screen "0890_Consumption" 1280x800, template "Navigation"
   on GenerateScreen: SetTag("DB_Zaehler_Anzeige_ReadWriteDeviceNo", 1); "Consumtion"(); SetBit("DB_Zaehler_Anzeige_Read"); function_b431313b(2, U 1, N); SetTag("Recipe_Appearance_Control", 4)
   IOField "Cumulative" at 366,244 size 100x30; FormatPattern 999999
      ProcessValue <- "DB_Zaehler_Anzeige_Gesamt_Anzahl"
   IOField "I/O field_2" at 473,244 size 170x30; FormatPattern 999999.99
      ProcessValue <- "DB_Zaehler_Anzeige_Gesamt_Verbrauch_K1"
      Visibility <- "DB790_PlantParameter_AmountMeteringUnits"
   IOField "I/O field_3" at 650,244 size 170x30; FormatPattern 999999.99
      ProcessValue <- "DB_Zaehler_Anzeige_Gesamt_Verbrauch_K2"
      Visibility <- "DB790_PlantParameter_AmountMeteringUnits"
   Button "Button_1" at 960,145 size 181x53; TextOff 'Last Shift'; TextOn 'Actual Shift'; TextList "Consumtion_Button"
      on Press: InvertBit("DB_Zaehler_Anzeige_ViewPreShift"); SetBit("DB_Zaehler_Anzeige_Read")
      ProcessValue <- "DB_Zaehler_Anzeige_ViewPreShift"
   IOField "I/O field_4" at 650,328 size 170x30; FormatPattern 999999.99
      ProcessValue <- "DB_Zaehler_Anzeige_Counter{1}_Verbrauch_K2"
      Visibility <- "DB790_PlantParameter_AmountMeteringUnits"
   IOField "I/O field_5" at 650,367 size 170x30; FormatPattern 999999.99
      ProcessValue <- "DB_Zaehler_Anzeige_Counter{2}_Verbrauch_K2"
      Visibility <- "DB790_PlantParameter_AmountMeteringUnits"
   IOField "I/O field_6" at 650,405 size 170x30; FormatPattern 999999.99
      ProcessValue <- "DB_Zaehler_Anzeige_Counter{3}_Verbrauch_K2"
      Visibility <- "DB790_PlantParameter_AmountMeteringUnits"
   IOField "I/O field_7" at 650,444 size 170x30; FormatPattern 999999.99
      ProcessValue <- "DB_Zaehler_Anzeige_Counter{4}_Verbrauch_K2"
      Visibility <- "DB790_PlantParameter_AmountMeteringUnits"
   IOField "I/O field_8" at 650,483 size 170x30; FormatPattern 999999.99
      ProcessValue <- "DB_Zaehler_Anzeige_Counter{5}_Verbrauch_K2"
      Visibility <- "DB790_PlantParameter_AmountMeteringUnits"
   IOField "I/O field_9" at 650,521 size 170x30; FormatPattern 999999.99
      ProcessValue <- "DB_Zaehler_Anzeige_Counter{6}_Verbrauch_K2"
      Visibility <- "DB790_PlantParameter_AmountMeteringUnits"
   IOField "I/O field_10" at 650,560 size 170x30; FormatPattern 999999.99
      ProcessValue <- "DB_Zaehler_Anzeige_Counter{7}_Verbrauch_K2"
      Visibility <- "DB790_PlantParameter_AmountMeteringUnits"
   IOField "I/O field_11" at 650,598 size 170x30; FormatPattern 999999.99
      ProcessValue <- "DB_Zaehler_Anzeige_Counter{8}_Verbrauch_K2"
      Visibility <- "DB790_PlantParameter_AmountMeteringUnits"
   IOField "I/O field_12" at 650,638 size 170x30; FormatPattern 999999.99
      ProcessValue <- "DB_Zaehler_Anzeige_Counter{9}_Verbrauch_K2"
      Visibility <- "DB790_PlantParameter_AmountMeteringUnits"
   IOField "I/O field_13" at 650,675 size 170x30; FormatPattern 999999.99
      ProcessValue <- "DB_Zaehler_Anzeige_Counter{10}_Verbrauch_K2"
      Visibility <- "DB790_PlantParameter_AmountMeteringUnits"
   IOField "I/O field_14" at 473,328 size 170x30; FormatPattern 999999.99
      ProcessValue <- "DB_Zaehler_Anzeige_Counter{1}_Verbrauch_K1"
      Visibility <- "DB790_PlantParameter_AmountMeteringUnits"
   IOField "I/O field_15" at 473,367 size 170x30; FormatPattern 999999.99
      ProcessValue <- "DB_Zaehler_Anzeige_Counter{2}_Verbrauch_K1"
      Visibility <- "DB790_PlantParameter_AmountMeteringUnits"
   IOField "I/O field_16" at 473,405 size 170x30; FormatPattern 999999.99
      ProcessValue <- "DB_Zaehler_Anzeige_Counter{3}_Verbrauch_K1"
      Visibility <- "DB790_PlantParameter_AmountMeteringUnits"
   IOField "I/O field_17" at 473,444 size 170x30; FormatPattern 999999.99
      ProcessValue <- "DB_Zaehler_Anzeige_Counter{4}_Verbrauch_K1"
      Visibility <- "DB790_PlantParameter_AmountMeteringUnits"
   IOField "I/O field_18" at 473,483 size 170x30; FormatPattern 999999.99
      ProcessValue <- "DB_Zaehler_Anzeige_Counter{5}_Verbrauch_K1"
      Visibility <- "DB790_PlantParameter_AmountMeteringUnits"
   IOField "I/O field_19" at 473,521 size 170x30; FormatPattern 999999.99
      ProcessValue <- "DB_Zaehler_Anzeige_Counter{6}_Verbrauch_K1"
      Visibility <- "DB790_PlantParameter_AmountMeteringUnits"
   IOField "I/O field_20" at 473,560 size 170x30; FormatPattern 999999.99
      ProcessValue <- "DB_Zaehler_Anzeige_Counter{7}_Verbrauch_K1"
      Visibility <- "DB790_PlantParameter_AmountMeteringUnits"
   IOField "I/O field_21" at 473,598 size 170x30; FormatPattern 999999.99
      ProcessValue <- "DB_Zaehler_Anzeige_Counter{8}_Verbrauch_K1"
      Visibility <- "DB790_PlantParameter_AmountMeteringUnits"
   IOField "I/O field_22" at 473,638 size 170x30; FormatPattern 999999.99
      ProcessValue <- "DB_Zaehler_Anzeige_Counter{9}_Verbrauch_K1"
      Visibility <- "DB790_PlantParameter_AmountMeteringUnits"
   IOField "I/O field_23" at 473,675 size 170x30; FormatPattern 999999.99
      ProcessValue <- "DB_Zaehler_Anzeige_Counter{10}_Verbrauch_K1"
      Visibility <- "DB790_PlantParameter_AmountMeteringUnits"
   IOField "I/O field_24" at 366,327 size 100x30; FormatPattern 999999
      ProcessValue <- "DB_Zaehler_Anzeige_Counter{1}_Anzahl"
   IOField "I/O field_25" at 366,365 size 100x30; FormatPattern 999999
      ProcessValue <- "DB_Zaehler_Anzeige_Counter{2}_Anzahl"
   IOField "I/O field_26" at 366,405 size 100x30; FormatPattern 999999
      ProcessValue <- "DB_Zaehler_Anzeige_Counter{3}_Anzahl"
   IOField "I/O field_27" at 366,443 size 100x30; FormatPattern 999999
      ProcessValue <- "DB_Zaehler_Anzeige_Counter{4}_Anzahl"
   IOField "I/O field_28" at 366,481 size 100x30; FormatPattern 999999
      ProcessValue <- "DB_Zaehler_Anzeige_Counter{5}_Anzahl"
   IOField "I/O field_29" at 366,520 size 100x30; FormatPattern 999999
      ProcessValue <- "DB_Zaehler_Anzeige_Counter{6}_Anzahl"
   IOField "I/O field_30" at 366,558 size 100x30; FormatPattern 999999
      ProcessValue <- "DB_Zaehler_Anzeige_Counter{7}_Anzahl"
   IOField "I/O field_31" at 366,598 size 100x30; FormatPattern 999999
      ProcessValue <- "DB_Zaehler_Anzeige_Counter{8}_Anzahl"
   IOField "I/O field_32" at 366,637 size 100x30; FormatPattern 999999
      ProcessValue <- "DB_Zaehler_Anzeige_Counter{9}_Anzahl"
   IOField "I/O field_33" at 365,676 size 100x30; FormatPattern 999999
      ProcessValue <- "DB_Zaehler_Anzeige_Counter{10}_Anzahl"
   IOField "I/O field_34" at 178,326 size 180x30; FormatPattern ????????????????????????????????????????????????????????????????????????????????
      ProcessValue <- "Consumtion_Name_1"
   IOField "I/O field_35" at 178,364 size 180x30; FormatPattern ????????????????????????????????????????????????????????????????????????????????
      ProcessValue <- "Consumtion_Name_2"
   IOField "I/O field_36" at 178,404 size 180x30; FormatPattern ????????????????????????????????????????????????????????????????????????????????
      ProcessValue <- "Consumtion_Name_3"
   IOField "I/O field_37" at 178,441 size 180x30; FormatPattern ????????????????????????????????????????????????????????????????????????????????
      ProcessValue <- "Consumtion_Name_4"
   IOField "I/O field_38" at 178,480 size 180x30; FormatPattern ????????????????????????????????????????????????????????????????????????????????
      ProcessValue <- "Consumtion_Name_5"
   IOField "I/O field_39" at 178,519 size 180x30; FormatPattern ????????????????????????????????????????????????????????????????????????????????
      ProcessValue <- "Consumtion_Name_6"
   IOField "I/O field_40" at 178,558 size 180x30; FormatPattern ????????????????????????????????????????????????????????????????????????????????
      ProcessValue <- "Consumtion_Name_7"
   IOField "I/O field_41" at 178,597 size 180x30; FormatPattern ????????????????????????????????????????????????????????????????????????????????
      ProcessValue <- "Consumtion_Name_8"
   IOField "I/O field_42" at 178,636 size 180x30; FormatPattern ????????????????????????????????????????????????????????????????????????????????
      ProcessValue <- "Consumtion_Name_9"
   IOField "I/O field_43" at 178,676 size 180x30; FormatPattern ????????????????????????????????????????????????????????????????????????????????
      ProcessValue <- "Consumtion_Name_10"
   Button "Button_3" at 326,99 size 451x32; TextOff 'Consumption'
   Button "Button_2" at 293,154 size 313x35; TextOff '001--010'; TextList "Consumtion"
      ProcessValue <- "DB_Zaehler_Anzeige_ReadWriteDeviceNo"
   Button "Button_6" at 650,280 size 170x30; TextOff '[KG]'
      Visibility <- "DB790_PlantParameter_AmountMeteringUnits"
   Button "Button_7" at 366,280 size 100x30; TextOff 'Amount'
   Button "Button_8" at 178,244 size 180x30; TextOff 'Cumulative'
   Button "Button_9" at 178,280 size 180x30; TextOff 'Name'
   Button "Button_10" at 111,280 size 60x30; TextOff 'No'
   Button "Button_11" at 473,280 size 170x30; TextOff '[KG]'
      Visibility <- "DB790_PlantParameter_AmountMeteringUnits"
   Button "Button_12" at 121,326 size 50x30; TextOff '.'
   Button "Button_13" at 121,364 size 50x30; TextOff '.'
   Button "Button_14" at 121,404 size 50x30; TextOff '.'
   Button "Button_15" at 121,441 size 50x30; TextOff '.'
   Button "Button_16" at 121,480 size 50x30; TextOff '.'
   Button "Button_17" at 121,519 size 50x30; TextOff '.'
   Button "Button_18" at 121,558 size 50x30; TextOff '.'
   Button "Button_19" at 121,597 size 50x30; TextOff '.'
   Button "Button_20" at 121,636 size 50x30; TextOff '.'
   Button "Button_21" at 121,676 size 50x30; TextOff '.'
   Button "b_incress_consumtion" at 618,154 size 46x35; TextOff 'Text'; PictureOff "NEXT"
      on Click: "Consumtion_Increase"(); "Consumtion"(); SetBit("DB_Zaehler_Anzeige_Read"); function_dd21b452("Consumtion Name Multiplexing Control", 1)
   Button "b_Decres_consumtion" at 234,154 size 46x35; TextOff 'Text'; PictureOff "BEFORE"
      on Click: "Consumtiom_Decrease"(); "Consumtion"(); SetBit("DB_Zaehler_Anzeige_Read"); function_b9b71300("Consumtion Name Multiplexing Control", 1)
   IOField "I/O field_44" at 473,208 size 170x30; FormatPattern ????????????????????
      ProcessValue <- "DB753_MeteringPump_Pump{1}_Name"
      Appearance <- "DB702_Tank_Value_Tank{1}_Color"
      Visibility <- "DB790_PlantParameter_AmountMeteringUnits"
   IOField "I/O field_45" at 650,208 size 170x30; FormatPattern ????????????????????
      ProcessValue <- "DB753_MeteringPump_Pump{2}_Name"
      Appearance <- "DB702_Tank_Value_Tank{2}_Color"
      Visibility <- "DB790_PlantParameter_AmountMeteringUnits"
   IOField "I/O field_46" at 826,244 size 170x30; FormatPattern 999999.99
      ProcessValue <- "DB_Zaehler_Anzeige_Gesamt_Verbrauch_K3"
      Visibility <- "DB790_PlantParameter_AmountMeteringUnits"
   IOField "I/O field_47" at 1001,244 size 170x30; FormatPattern 999999.99
      ProcessValue <- "DB_Zaehler_Anzeige_Gesamt_Verbrauch_K4"
      Visibility <- "DB790_PlantParameter_AmountMeteringUnits"
   IOField "I/O field_48" at 1001,328 size 170x30; FormatPattern 999999.99
      ProcessValue <- "DB_Zaehler_Anzeige_Counter{1}_Verbrauch_K4"
      Visibility <- "DB790_PlantParameter_AmountMeteringUnits"
   IOField "I/O field_49" at 1001,367 size 170x30; FormatPattern 999999.99
      ProcessValue <- "DB_Zaehler_Anzeige_Counter{2}_Verbrauch_K4"
      Visibility <- "DB790_PlantParameter_AmountMeteringUnits"
   IOField "I/O field_50" at 1001,405 size 170x30; FormatPattern 999999.99
      ProcessValue <- "DB_Zaehler_Anzeige_Counter{3}_Verbrauch_K4"
      Visibility <- "DB790_PlantParameter_AmountMeteringUnits"
   IOField "I/O field_51" at 1001,444 size 170x30; FormatPattern 999999.99
      ProcessValue <- "DB_Zaehler_Anzeige_Counter{4}_Verbrauch_K4"
      Visibility <- "DB790_PlantParameter_AmountMeteringUnits"
   IOField "I/O field_52" at 1001,483 size 170x30; FormatPattern 999999.99
      ProcessValue <- "DB_Zaehler_Anzeige_Counter{5}_Verbrauch_K4"
      Visibility <- "DB790_PlantParameter_AmountMeteringUnits"
   IOField "I/O field_53" at 1001,521 size 170x30; FormatPattern 999999.99
      ProcessValue <- "DB_Zaehler_Anzeige_Counter{6}_Verbrauch_K4"
      Visibility <- "DB790_PlantParameter_AmountMeteringUnits"
   IOField "I/O field_54" at 1001,560 size 170x30; FormatPattern 999999.99
      ProcessValue <- "DB_Zaehler_Anzeige_Counter{7}_Verbrauch_K4"
      Visibility <- "DB790_PlantParameter_AmountMeteringUnits"
   IOField "I/O field_55" at 1001,598 size 170x30; FormatPattern 999999.99
      ProcessValue <- "DB_Zaehler_Anzeige_Counter{8}_Verbrauch_K4"
      Visibility <- "DB790_PlantParameter_AmountMeteringUnits"
   IOField "I/O field_56" at 1001,638 size 170x30; FormatPattern 999999.99
      ProcessValue <- "DB_Zaehler_Anzeige_Counter{9}_Verbrauch_K4"
      Visibility <- "DB790_PlantParameter_AmountMeteringUnits"
   IOField "I/O field_57" at 1001,675 size 170x30; FormatPattern 999999.99
      ProcessValue <- "DB_Zaehler_Anzeige_Counter{10}_Verbrauch_K4"
      Visibility <- "DB790_PlantParameter_AmountMeteringUnits"
   IOField "I/O field_58" at 826,328 size 170x30; FormatPattern 999999.99
      ProcessValue <- "DB_Zaehler_Anzeige_Counter{1}_Verbrauch_K3"
      Visibility <- "DB790_PlantParameter_AmountMeteringUnits"
   IOField "I/O field_59" at 826,367 size 170x30; FormatPattern 999999.99
      ProcessValue <- "DB_Zaehler_Anzeige_Counter{2}_Verbrauch_K3"
      Visibility <- "DB790_PlantParameter_AmountMeteringUnits"
   IOField "I/O field_60" at 826,405 size 170x30; FormatPattern 999999.99
      ProcessValue <- "DB_Zaehler_Anzeige_Counter{3}_Verbrauch_K3"
      Visibility <- "DB790_PlantParameter_AmountMeteringUnits"
   IOField "I/O field_61" at 826,444 size 170x30; FormatPattern 999999.99
      ProcessValue <- "DB_Zaehler_Anzeige_Counter{4}_Verbrauch_K3"
      Visibility <- "DB790_PlantParameter_AmountMeteringUnits"
   IOField "I/O field_62" at 826,483 size 170x30; FormatPattern 999999.99
      ProcessValue <- "DB_Zaehler_Anzeige_Counter{5}_Verbrauch_K3"
      Visibility <- "DB790_PlantParameter_AmountMeteringUnits"
   IOField "I/O field_63" at 826,521 size 170x30; FormatPattern 999999.99
      ProcessValue <- "DB_Zaehler_Anzeige_Counter{6}_Verbrauch_K3"
      Visibility <- "DB790_PlantParameter_AmountMeteringUnits"
   IOField "I/O field_64" at 826,560 size 170x30; FormatPattern 999999.99
      ProcessValue <- "DB_Zaehler_Anzeige_Counter{7}_Verbrauch_K3"
      Visibility <- "DB790_PlantParameter_AmountMeteringUnits"
   IOField "I/O field_65" at 826,598 size 170x30; FormatPattern 999999.99
      ProcessValue <- "DB_Zaehler_Anzeige_Counter{8}_Verbrauch_K3"
      Visibility <- "DB790_PlantParameter_AmountMeteringUnits"
   IOField "I/O field_66" at 826,638 size 170x30; FormatPattern 999999.99
      ProcessValue <- "DB_Zaehler_Anzeige_Counter{9}_Verbrauch_K3"
      Visibility <- "DB790_PlantParameter_AmountMeteringUnits"
   IOField "I/O field_67" at 826,675 size 170x30; FormatPattern 999999.99
      ProcessValue <- "DB_Zaehler_Anzeige_Counter{10}_Verbrauch_K3"
      Visibility <- "DB790_PlantParameter_AmountMeteringUnits"
   Button "Button_4" at 1001,280 size 170x30; TextOff '[KG]'
      Visibility <- "DB790_PlantParameter_AmountMeteringUnits"
   Button "Button_5" at 826,280 size 170x30; TextOff '[KG]'
      Visibility <- "DB790_PlantParameter_AmountMeteringUnits"
   IOField "I/O field_68" at 826,208 size 170x30; FormatPattern ????????????????????
      ProcessValue <- "DB753_MeteringPump_Pump{3}_Name"
      Visibility <- "DB790_PlantParameter_AmountMeteringUnits"
      Appearance <- "DB702_Tank_Value_Tank{3}_Color"
   IOField "I/O field_69" at 1001,208 size 170x30; FormatPattern ????????????????????
      ProcessValue <- "DB753_MeteringPump_Pump{4}_Name"
      Visibility <- "DB790_PlantParameter_AmountMeteringUnits"
      Appearance <- "DB702_Tank_Value_Tank{4}_Color"
   Button "b_ShifProto_ShotCounter_1" at 208,713 size 60x60; TextOff 'Shot Counter'; PictureList "ico_ShiftProtocol"
      ProcessValue <- "Recipe_Appearance_Control"
      Appearance <- "Recipe_Appearance_Control"
   Button "b_Shiftproto_shiftproto" at 208,713 size 60x60; TextOff 'Shift proto'
      on Click: ActivateScreen("0112_Shift protocol", 0); SetTag("Recipe_Appearance_Control", 2)
      Appearance <- "Recipe_Appearance_Control"
   Button "b_SC" at 478,713 size 60x60; TextOff 'Shot Counter'; PictureList "ico_ShotCounter"
      on Press: ActivateScreen("0891_Shotcounter MixingHead", 0); SetTag("Recipe_Appearance_Control", 5)
      Appearance <- "Recipe_Appearance_Control"
      ProcessValue <- "Recipe_Appearance_Control"
   Button "b_SC_1" at 478,713 size 60x60; TextOff 'Shot Counter'
      on Click: ActivateScreen("0891_Shotcounter MixingHead", 0); SetTag("Recipe_Appearance_Control", 5)
      Appearance <- "Recipe_Appearance_Control"
   Button "b_Shift_Plan" at 118,713 size 60x60; TextOff 'Shift Plan'; PictureList "ico_ShiftPlan"
      on Press: ActivateScreen("0113_SettingShiftPlan", 0); SetTag("Recipe_Appearance_Control", 1)
      Appearance <- "Recipe_Appearance_Control"
      ProcessValue <- "Recipe_Appearance_Control"
   Button "b_Shift_Plan_1" at 118,713 size 60x60; TextOff 'Shift Plan'
      on Click: "SettingShiftPlan"(); ActivateScreen("0113_SettingShiftPlan", 0); SetTag("Recipe_Appearance_Control", 1)
      Appearance <- "Recipe_Appearance_Control"
   Button "b_LS_Lastshot" at 298,713 size 60x60; TextOff 'Last Shot'; PictureList "ico_LastShot"
      on Press: ActivateScreen("0036_Last Shot", 0); SetTag("Recipe_Appearance_Control", 3)
      Appearance <- "Recipe_Appearance_Control"
      ProcessValue <- "Recipe_Appearance_Control"
   Button "b_LS_Lastshot_1" at 298,713 size 60x60; TextOff 'Last Shot'
      on Click: ActivateScreen("0036_Last Shot", 0); SetTag("Recipe_Appearance_Control", 3)
      Appearance <- "Recipe_Appearance_Control"
   Button "b_Consumtion" at 388,713 size 60x60; TextOff 'Consumtion / Consum'; PictureList "ico_consum"
      on Press: ActivateScreen("0890_Consumption", 0); SetTag("Recipe_Appearance_Control", 4)
      Appearance <- "Recipe_Appearance_Control"
      ProcessValue <- "Recipe_Appearance_Control"
   Button "b_Consumtion_1" at 388,713 size 60x60; TextOff 'Consumtion / Consum'
      on Click: ActivateScreen("0890_Consumption", 0); SetTag("Recipe_Appearance_Control", 4)
      Appearance <- "Recipe_Appearance_Control"

screen "0891_Shotcounter MixingHead" 1280x800, template "Navigation"
   on GenerateScreen: SetBit("DB_Zaehler_Anzeige_Read"); SetTag("Recipe_Appearance_Control", 5)
   IOField "I/O field_14" at 378,202 size 168x30; FormatPattern 9999999
      ProcessValue <- "DB_Zaehler_Anzeige_MH_Counter_ActualShift{1}"
      Visibility <- "DB790_PlantParameter_AmountMH"
   IOField "lastshift1" at 564,202 size 168x30; FormatPattern 9999999
      ProcessValue <- "DB_Zaehler_Anzeige_MH_Counter_PreShift{1}"
      Visibility <- "DB790_PlantParameter_AmountMH"
   IOField "I/O field_2" at 748,202 size 168x30; Authorization "User administration"; FormatPattern 9999999
      ProcessValue <- "DB_Zaehler_Anzeige_MH_Counter_Reset{1}"
      Visibility <- "DB790_PlantParameter_AmountMH"
   IOField "I/O field_3" at 933,202 size 168x30; FormatPattern 9999999
      ProcessValue <- "DB_Zaehler_Anzeige_MH_Counter_NonReset{1}"
      Visibility <- "DB790_PlantParameter_AmountMH"
   Button "Button_3" at 326,104 size 451x32; TextOff 'Shot counter Mixinghead'
   Button "Button_1" at 378,158 size 168x30; TextOff 'Actual Shift'
   Button "Button_2" at 564,158 size 168x30; TextOff 'Last Shift'
   Button "Button_4" at 748,158 size 168x30; TextOff 'Resetable'
   Button "Button_5" at 933,158 size 168x30; TextOff 'Cumulative'
   Button "Button_6" at 309,202 size 50x30; TextOff '1.'
      Visibility <- "DB790_PlantParameter_AmountMH"
   IOField "I/O field_4" at 378,245 size 168x30; FormatPattern 9999999
      ProcessValue <- "DB_Zaehler_Anzeige_MH_Counter_ActualShift{2}"
      Visibility <- "DB790_PlantParameter_AmountMH"
   IOField "I/O field_5" at 564,245 size 168x30; FormatPattern 9999999
      ProcessValue <- "DB_Zaehler_Anzeige_MH_Counter_PreShift{2}"
      Visibility <- "DB790_PlantParameter_AmountMH"
   IOField "I/O field_6" at 748,245 size 168x30; Authorization "User administration"; FormatPattern 9999999
      ProcessValue <- "DB_Zaehler_Anzeige_MH_Counter_Reset{2}"
      Visibility <- "DB790_PlantParameter_AmountMH"
   IOField "I/O field_7" at 933,245 size 168x30; FormatPattern 9999999
      ProcessValue <- "DB_Zaehler_Anzeige_MH_Counter_NonReset{2}"
      Visibility <- "DB790_PlantParameter_AmountMH"
   Button "Button_7" at 309,245 size 50x30; TextOff '2.'
      Visibility <- "DB790_PlantParameter_AmountMH"
   IOField "I/O field_8" at 378,290 size 168x30; FormatPattern 9999999
      ProcessValue <- "DB_Zaehler_Anzeige_MH_Counter_ActualShift{3}"
      Visibility <- "DB790_PlantParameter_AmountMH"
   IOField "I/O field_9" at 564,290 size 168x30; FormatPattern 9999999
      ProcessValue <- "DB_Zaehler_Anzeige_MH_Counter_PreShift{3}"
      Visibility <- "DB790_PlantParameter_AmountMH"
   IOField "I/O field_10" at 748,290 size 168x30; Authorization "User administration"; FormatPattern 9999999
      ProcessValue <- "DB_Zaehler_Anzeige_MH_Counter_Reset{3}"
      Visibility <- "DB790_PlantParameter_AmountMH"
   IOField "I/O field_11" at 933,290 size 168x30; FormatPattern 9999999
      ProcessValue <- "DB_Zaehler_Anzeige_MH_Counter_NonReset{3}"
      Visibility <- "DB790_PlantParameter_AmountMH"
   Button "Button_8" at 309,290 size 50x30; TextOff '3.'
      Visibility <- "DB790_PlantParameter_AmountMH"
   IOField "I/O field_12" at 378,334 size 168x30; FormatPattern 9999999
      ProcessValue <- "DB_Zaehler_Anzeige_MH_Counter_ActualShift{4}"
      Visibility <- "DB790_PlantParameter_AmountMH"
   IOField "I/O field_13" at 564,334 size 168x30; FormatPattern 9999999
      ProcessValue <- "DB_Zaehler_Anzeige_MH_Counter_PreShift{4}"
      Visibility <- "DB790_PlantParameter_AmountMH"
   IOField "I/O field_15" at 748,334 size 168x30; Authorization "User administration"; FormatPattern 9999999
      ProcessValue <- "DB_Zaehler_Anzeige_MH_Counter_Reset{4}"
      Visibility <- "DB790_PlantParameter_AmountMH"
   IOField "I/O field_16" at 933,334 size 168x30; FormatPattern 9999999
      ProcessValue <- "DB_Zaehler_Anzeige_MH_Counter_NonReset{4}"
      Visibility <- "DB790_PlantParameter_AmountMH"
   Button "Button_9" at 309,334 size 50x30; TextOff '4.'
      Visibility <- "DB790_PlantParameter_AmountMH"
   IOField "I/O field_17" at 378,378 size 168x30; FormatPattern 9999999
      ProcessValue <- "DB_Zaehler_Anzeige_MH_Counter_ActualShift{5}"
      Visibility <- "DB790_PlantParameter_AmountMH"
   IOField "I/O field_18" at 564,378 size 168x30; FormatPattern 9999999
      ProcessValue <- "DB_Zaehler_Anzeige_MH_Counter_PreShift{5}"
      Visibility <- "DB790_PlantParameter_AmountMH"
   IOField "I/O field_19" at 748,378 size 168x30; Authorization "User administration"; FormatPattern 9999999
      ProcessValue <- "DB_Zaehler_Anzeige_MH_Counter_Reset{5}"
      Visibility <- "DB790_PlantParameter_AmountMH"
   IOField "I/O field_20" at 933,378 size 168x30; FormatPattern 9999999
      ProcessValue <- "DB_Zaehler_Anzeige_MH_Counter_NonReset{5}"
      Visibility <- "DB790_PlantParameter_AmountMH"
   Button "Button_10" at 309,378 size 50x30; TextOff '5.'
      Visibility <- "DB790_PlantParameter_AmountMH"
   IOField "I/O field_21" at 378,421 size 168x30; FormatPattern 9999999
      ProcessValue <- "DB_Zaehler_Anzeige_MH_Counter_ActualShift{6}"
      Visibility <- "DB790_PlantParameter_AmountMH"
   IOField "I/O field_22" at 564,421 size 168x30; FormatPattern 9999999
      ProcessValue <- "DB_Zaehler_Anzeige_MH_Counter_PreShift{6}"
      Visibility <- "DB790_PlantParameter_AmountMH"
   IOField "I/O field_23" at 748,421 size 168x30; Authorization "User administration"; FormatPattern 9999999
      ProcessValue <- "DB_Zaehler_Anzeige_MH_Counter_Reset{6}"
      Visibility <- "DB790_PlantParameter_AmountMH"
   IOField "I/O field_24" at 933,421 size 168x30; FormatPattern 9999999
      ProcessValue <- "DB_Zaehler_Anzeige_MH_Counter_NonReset{6}"
      Visibility <- "DB790_PlantParameter_AmountMH"
   Button "Button_11" at 309,421 size 50x30; TextOff '6.'
      Visibility <- "DB790_PlantParameter_AmountMH"
   IOField "I/O field_25" at 378,464 size 168x30; FormatPattern 9999999
      ProcessValue <- "DB_Zaehler_Anzeige_MH_Counter_ActualShift{7}"
      Visibility <- "DB790_PlantParameter_AmountMH"
   IOField "I/O field_26" at 564,464 size 168x30; FormatPattern 9999999
      ProcessValue <- "DB_Zaehler_Anzeige_MH_Counter_PreShift{7}"
      Visibility <- "DB790_PlantParameter_AmountMH"
   IOField "I/O field_27" at 748,464 size 168x30; Authorization "User administration"; FormatPattern 9999999
      ProcessValue <- "DB_Zaehler_Anzeige_MH_Counter_Reset{7}"
      Visibility <- "DB790_PlantParameter_AmountMH"
   IOField "I/O field_28" at 933,464 size 168x30; FormatPattern 9999999
      ProcessValue <- "DB_Zaehler_Anzeige_MH_Counter_NonReset{7}"
      Visibility <- "DB790_PlantParameter_AmountMH"
   Button "Button_12" at 309,464 size 50x30; TextOff '7.'
      Visibility <- "DB790_PlantParameter_AmountMH"
   IOField "I/O field_29" at 378,507 size 168x30; FormatPattern 9999999
      ProcessValue <- "DB_Zaehler_Anzeige_MH_Counter_ActualShift{8}"
      Visibility <- "DB790_PlantParameter_AmountMH"
   IOField "I/O field_30" at 564,507 size 168x30; FormatPattern 9999999
      ProcessValue <- "DB_Zaehler_Anzeige_MH_Counter_PreShift{8}"
      Visibility <- "DB790_PlantParameter_AmountMH"
   IOField "I/O field_31" at 748,507 size 168x30; Authorization "User administration"; FormatPattern 9999999
      ProcessValue <- "DB_Zaehler_Anzeige_MH_Counter_Reset{8}"
      Visibility <- "DB790_PlantParameter_AmountMH"
   IOField "I/O field_32" at 933,507 size 168x30; FormatPattern 9999999
      ProcessValue <- "DB_Zaehler_Anzeige_MH_Counter_NonReset{8}"
      Visibility <- "DB790_PlantParameter_AmountMH"
   Button "Button_13" at 309,507 size 50x30; TextOff '8.'
      Visibility <- "DB790_PlantParameter_AmountMH"
   IOField "I/O field_33" at 378,551 size 168x30; FormatPattern 9999999
      ProcessValue <- "DB_Zaehler_Anzeige_MH_Counter_ActualShift{9}"
      Visibility <- "DB790_PlantParameter_AmountMH"
   IOField "I/O field_34" at 564,551 size 168x30; FormatPattern 9999999
      ProcessValue <- "DB_Zaehler_Anzeige_MH_Counter_PreShift{9}"
      Visibility <- "DB790_PlantParameter_AmountMH"
   IOField "I/O field_35" at 748,551 size 168x30; Authorization "User administration"; FormatPattern 9999999
      ProcessValue <- "DB_Zaehler_Anzeige_MH_Counter_Reset{9}"
      Visibility <- "DB790_PlantParameter_AmountMH"
   IOField "I/O field_36" at 933,551 size 168x30; FormatPattern 9999999
      ProcessValue <- "DB_Zaehler_Anzeige_MH_Counter_NonReset{9}"
      Visibility <- "DB790_PlantParameter_AmountMH"
   Button "Button_14" at 309,551 size 50x30; TextOff '9.'
      Visibility <- "DB790_PlantParameter_AmountMH"
   IOField "I/O field_37" at 378,594 size 168x30; FormatPattern 9999999
      ProcessValue <- "DB_Zaehler_Anzeige_MH_Counter_ActualShift{10}"
      Visibility <- "DB790_PlantParameter_AmountMH"
   IOField "I/O field_38" at 564,594 size 168x30; FormatPattern 9999999
      ProcessValue <- "DB_Zaehler_Anzeige_MH_Counter_PreShift{10}"
      Visibility <- "DB790_PlantParameter_AmountMH"
   IOField "I/O field_39" at 748,594 size 168x30; Authorization "User administration"; FormatPattern 9999999
      ProcessValue <- "DB_Zaehler_Anzeige_MH_Counter_Reset{10}"
      Visibility <- "DB790_PlantParameter_AmountMH"
   IOField "I/O field_40" at 933,594 size 168x30; FormatPattern 9999999
      ProcessValue <- "DB_Zaehler_Anzeige_MH_Counter_NonReset{10}"
      Visibility <- "DB790_PlantParameter_AmountMH"
   Button "Button_15" at 309,594 size 50x30; TextOff '10.'
      Visibility <- "DB790_PlantParameter_AmountMH"
   GraphicView "Graphic view_3" at 108,290 size 177x240; Picture "images_4"
   Button "b_ShifProto_ShotCounter_1" at 208,713 size 60x60; TextOff 'Shot Counter'; PictureList "ico_ShiftProtocol"
      ProcessValue <- "Recipe_Appearance_Control"
      Appearance <- "Recipe_Appearance_Control"
   Button "b_Shiftproto_shiftproto" at 208,713 size 60x60; TextOff 'Shift proto'
      on Click: ActivateScreen("0112_Shift protocol", 0); SetTag("Recipe_Appearance_Control", 2)
      Appearance <- "Recipe_Appearance_Control"
   Button "b_SC" at 478,713 size 60x60; TextOff 'Shot Counter'; PictureList "ico_ShotCounter"
      on Press: ActivateScreen("0891_Shotcounter MixingHead", 0); SetTag("Recipe_Appearance_Control", 5)
      Appearance <- "Recipe_Appearance_Control"
      ProcessValue <- "Recipe_Appearance_Control"
   Button "b_SC_1" at 478,713 size 60x60; TextOff 'Shot Counter'
      on Click: ActivateScreen("0891_Shotcounter MixingHead", 0); SetTag("Recipe_Appearance_Control", 5)
      Appearance <- "Recipe_Appearance_Control"
   Button "b_Shift_Plan" at 118,713 size 60x60; TextOff 'Shift Plan'; PictureList "ico_ShiftPlan"
      on Press: ActivateScreen("0113_SettingShiftPlan", 0); SetTag("Recipe_Appearance_Control", 1)
      Appearance <- "Recipe_Appearance_Control"
      ProcessValue <- "Recipe_Appearance_Control"
   Button "b_Shift_Plan_1" at 118,713 size 60x60; TextOff 'Shift Plan'
      on Click: "SettingShiftPlan"(); ActivateScreen("0113_SettingShiftPlan", 0); SetTag("Recipe_Appearance_Control", 1)
      Appearance <- "Recipe_Appearance_Control"
   Button "b_LS_Lastshot" at 298,713 size 60x60; TextOff 'Last Shot'; PictureList "ico_LastShot"
      on Press: ActivateScreen("0036_Last Shot", 0); SetTag("Recipe_Appearance_Control", 3)
      Appearance <- "Recipe_Appearance_Control"
      ProcessValue <- "Recipe_Appearance_Control"
   Button "b_LS_Lastshot_1" at 298,713 size 60x60; TextOff 'Last Shot'
      on Click: ActivateScreen("0036_Last Shot", 0); SetTag("Recipe_Appearance_Control", 3)
      Appearance <- "Recipe_Appearance_Control"
   Button "b_Consumtion" at 388,713 size 60x60; TextOff 'Consumtion / Consum'; PictureList "ico_consum"
      on Press: ActivateScreen("0890_Consumption", 0); SetTag("Recipe_Appearance_Control", 4)
      Appearance <- "Recipe_Appearance_Control"
      ProcessValue <- "Recipe_Appearance_Control"
   Button "b_Consumtion_1" at 388,713 size 60x60; TextOff 'Consumtion / Consum'
      on Click: ActivateScreen("0890_Consumption", 0); SetTag("Recipe_Appearance_Control", 4)
      Appearance <- "Recipe_Appearance_Control"

screen "0892_Tool Editor" 1280x800, template "Navigation"
   on GenerateScreen: SetTag("InterfaceVisu_ReadWriteDeviceNo", "DB_MouldEditor_HMI_uData_sSelected_iTool"); SetTag("DB_MouldEditor_HMI_uData_sSelected_sPS_iPS", 1); SetTag("NavScreenChange", 6)
   on ClearScreen: SetTag("NavScreenChange", 0)
   Rectangle "Rectangle_3" at 346,760 size 73x12
      Visibility <- "DB704_MH_Value_Mixinghead{0}_AmountComponent"
   Rectangle "Rectangle_5" at 482,760 size 73x12
      Visibility <- "DB704_MH_Value_Mixinghead{0}_AmountComponent"
   Rectangle "Rectangle_9" at 617,760 size 73x12
      Visibility <- "DB704_MH_Value_Mixinghead{0}_AmountComponent"
   Rectangle "Rectangle_10" at 751,760 size 73x12
      Visibility <- "DB704_MH_Value_Mixinghead{0}_AmountComponent"
   Rectangle "Rectangle_14" at 887,760 size 73x12
      Visibility <- "DB704_MH_Value_Mixinghead{0}_AmountComponent"
   Rectangle "Rectangle_15" at 1024,760 size 73x12
      Visibility <- "DB704_MH_Value_Mixinghead{0}_AmountComponent"
   Button "Button_40" at 994,502 size 66x32; TextOff 'Text'
      Visibility <- "DB_MouldEditor_HMI_uData_uTools_PartShot_Amount"
      Appearance <- "DB_MouldEditor_HMI_uData_sSelected_sPS_iPS"
   Button "Button_39" at 928,502 size 66x32; TextOff 'Text'
      Visibility <- "DB_MouldEditor_HMI_uData_uTools_PartShot_Amount"
      Appearance <- "DB_MouldEditor_HMI_uData_sSelected_sPS_iPS"
   Button "Button_38" at 852,502 size 75x32; TextOff 'Text'
      Visibility <- "DB_MouldEditor_HMI_uData_uTools_PartShot_Amount"
      Appearance <- "DB_MouldEditor_HMI_uData_sSelected_sPS_iPS"
   Button "Button_37" at 994,467 size 66x32; TextOff 'Text'
      Visibility <- "DB_MouldEditor_HMI_uData_uTools_PartShot_Amount"
      Appearance <- "DB_MouldEditor_HMI_uData_sSelected_sPS_iPS"
   Button "Button_36" at 928,467 size 66x32; TextOff 'Text'
      Visibility <- "DB_MouldEditor_HMI_uData_uTools_PartShot_Amount"
      Appearance <- "DB_MouldEditor_HMI_uData_sSelected_sPS_iPS"
   Button "Button_35" at 852,467 size 75x32; TextOff 'Text'
      Visibility <- "DB_MouldEditor_HMI_uData_uTools_PartShot_Amount"
      Appearance <- "DB_MouldEditor_HMI_uData_sSelected_sPS_iPS"
   Button "Button_34" at 994,432 size 66x32; TextOff 'Text'
      Visibility <- "DB_MouldEditor_HMI_uData_uTools_PartShot_Amount"
      Appearance <- "DB_MouldEditor_HMI_uData_sSelected_sPS_iPS"
   Button "Button_33" at 928,432 size 66x32; TextOff 'Text'
      Visibility <- "DB_MouldEditor_HMI_uData_uTools_PartShot_Amount"
      Appearance <- "DB_MouldEditor_HMI_uData_sSelected_sPS_iPS"
   Button "Button_32" at 852,432 size 75x32; TextOff 'Text'
      Visibility <- "DB_MouldEditor_HMI_uData_uTools_PartShot_Amount"
      Appearance <- "DB_MouldEditor_HMI_uData_sSelected_sPS_iPS"
   Button "Button_31" at 994,397 size 66x32; TextOff 'Text'
      Visibility <- "DB_MouldEditor_HMI_uData_uTools_PartShot_Amount"
      Appearance <- "DB_MouldEditor_HMI_uData_sSelected_sPS_iPS"
   Button "Button_30" at 928,397 size 66x32; TextOff 'Text'
      Visibility <- "DB_MouldEditor_HMI_uData_uTools_PartShot_Amount"
      Appearance <- "DB_MouldEditor_HMI_uData_sSelected_sPS_iPS"
   Button "Button_29" at 852,397 size 75x32; TextOff 'Text'
      Visibility <- "DB_MouldEditor_HMI_uData_uTools_PartShot_Amount"
      Appearance <- "DB_MouldEditor_HMI_uData_sSelected_sPS_iPS"
   Button "Button_28" at 994,362 size 66x32; TextOff 'Text'
      Visibility <- "DB_MouldEditor_HMI_uData_uTools_PartShot_Amount"
      Appearance <- "DB_MouldEditor_HMI_uData_sSelected_sPS_iPS"
   Button "Button_27" at 928,362 size 66x32; TextOff 'Text'
      Visibility <- "DB_MouldEditor_HMI_uData_uTools_PartShot_Amount"
      Appearance <- "DB_MouldEditor_HMI_uData_sSelected_sPS_iPS"
   Button "Button_26" at 852,362 size 75x32; TextOff 'Text'
      Visibility <- "DB_MouldEditor_HMI_uData_uTools_PartShot_Amount"
      Appearance <- "DB_MouldEditor_HMI_uData_sSelected_sPS_iPS"
   Button "Button_25" at 994,327 size 66x32; TextOff 'Text'
      Visibility <- "DB_MouldEditor_HMI_uData_uTools_PartShot_Amount"
      Appearance <- "DB_MouldEditor_HMI_uData_sSelected_sPS_iPS"
   Button "Button_24" at 928,327 size 66x32; TextOff 'Text'
      Visibility <- "DB_MouldEditor_HMI_uData_uTools_PartShot_Amount"
      Appearance <- "DB_MouldEditor_HMI_uData_sSelected_sPS_iPS"
   Button "Button_23" at 852,327 size 75x32; TextOff 'Text'
      Visibility <- "DB_MouldEditor_HMI_uData_uTools_PartShot_Amount"
      Appearance <- "DB_MouldEditor_HMI_uData_sSelected_sPS_iPS"
   Button "Button_22" at 994,293 size 66x32; TextOff 'Text'
      Visibility <- "DB_MouldEditor_HMI_uData_uTools_PartShot_Amount"
      Appearance <- "DB_MouldEditor_HMI_uData_sSelected_sPS_iPS"
   Button "Button_21" at 928,293 size 66x32; TextOff 'Text'
      Visibility <- "DB_MouldEditor_HMI_uData_uTools_PartShot_Amount"
      Appearance <- "DB_MouldEditor_HMI_uData_sSelected_sPS_iPS"
   Button "Button_20" at 852,293 size 75x32; TextOff 'Text'
      Visibility <- "DB_MouldEditor_HMI_uData_uTools_PartShot_Amount"
      Appearance <- "DB_MouldEditor_HMI_uData_sSelected_sPS_iPS"
   Button "Button_19" at 994,258 size 66x32; TextOff 'Text'
      Visibility <- "DB_MouldEditor_HMI_uData_uTools_PartShot_Amount"
      Appearance <- "DB_MouldEditor_HMI_uData_sSelected_sPS_iPS"
   Button "Button_18" at 928,258 size 66x32; TextOff 'Text'
      Visibility <- "DB_MouldEditor_HMI_uData_uTools_PartShot_Amount"
      Appearance <- "DB_MouldEditor_HMI_uData_sSelected_sPS_iPS"
   Button "Button_17" at 852,258 size 75x32; TextOff 'Text'
      Visibility <- "DB_MouldEditor_HMI_uData_uTools_PartShot_Amount"
      Appearance <- "DB_MouldEditor_HMI_uData_sSelected_sPS_iPS"
   TextField "Text field_1" at 141,143 size 208x35; Text 'Tool No :'
   IOField "itool" at 355,143 size 57x35; FormatPattern 999
      ProcessValue <- "DB_MouldEditor_HMI_uData_sSelected_iTool"
   TextField "Text field_2" at 465,143 size 200x35; Text 'Tool Name :'
      Visibility <- "DB_MouldEditor_HMI_uData_uTools_PartShot_Amount"
   IOField "I/O field_3" at 235,258 size 84x32; Authorization "Operate"; FormatPattern 999
      ProcessValue <- "DB_MouldEditor_HMI_uData_arShotSet{1}_MHNo"
      Visibility <- "DB_MouldEditor_HMI_uData_uTools_PartShot_Amount"
      Appearance <- "DB_MouldEditor_HMI_uData_sSelected_sPS_iPS"
   IOField "Shottime_1" at 318,258 size 150x32; Authorization "Operate"; FormatPattern 99.999
      ProcessValue <- "DB_MouldEditor_HMI_uData_arShotSet{1}_FoamingTime"
      Visibility <- "DB_MouldEditor_HMI_uData_uTools_PartShot_Amount"
      ObjectEnable <- "DB_MouldEditor_HMI_uData_sSelected_iCalculation"
      Appearance <- "DB_MouldEditor_HMI_uData_sSelected_sPS_iPS"
   IOField "totalflow_1" at 467,258 size 144x32; Authorization "Operate"; FormatPattern 9999.99
      ProcessValue <- "DB_MouldEditor_HMI_uData_sCalculatedValues_arTotalFlow{1}"
      Visibility <- "DB_MouldEditor_HMI_uData_uTools_PartShot_Amount"
      ObjectEnable <- "DB_MouldEditor_HMI_uData_sSelected_iCalculation"
      Appearance <- "DB_MouldEditor_HMI_uData_sSelected_sPS_iPS"
   IOField "totalweight_1" at 609,258 size 151x32; Authorization "Operate"; FormatPattern 999.99
      ProcessValue <- "DB_MouldEditor_HMI_uData_arShotSet{1}_PartWeight"
      Visibility <- "DB_MouldEditor_HMI_uData_uTools_PartShot_Amount"
      ObjectEnable <- "DB_MouldEditor_HMI_uData_sSelected_iCalculation"
      Appearance <- "DB_MouldEditor_HMI_uData_sSelected_sPS_iPS"
   IOField "I/O field_7" at 759,258 size 93x32; Authorization "Operate"; FormatPattern 9999
      ProcessValue <- "DB_MouldEditor_HMI_uData_arShotSet{1}_PartCounter"
      Visibility <- "DB_MouldEditor_HMI_uData_uTools_PartShot_Amount"
      Appearance <- "DB_MouldEditor_HMI_uData_sSelected_sPS_iPS"
   TextField "Text field_4" at 148,229 size 89x30; Text 'PS'
   TextField "Text field_5" at 235,229 size 84x30; Text 'MH'
   TextField "Text field_6" at 318,229 size 150x30; Text 'Shottime / Shot time'
      Appearance <- "DB_MouldEditor_HMI_uData_sSelected_iCalculation"
   TextField "Text field_7" at 467,229 size 144x30; Text 'total Flow'
      Appearance <- "DB_MouldEditor_HMI_uData_sSelected_iCalculation"
   TextField "Text field_8" at 609,229 size 151x30; Text 'total Weight'
      Appearance <- "DB_MouldEditor_HMI_uData_sSelected_iCalculation"
   TextField "Text field_9" at 759,229 size 95x30; Text 'Counter'
   TextField "Text field_10" at 852,229 size 79x30; Text 'Service'
   TextField "Text field_11" at 928,229 size 68x30; Text 'CP'
   Button "Button_1" at 517,585 size 120x33; TextOff 'Deactivate'; TextOn 'Activate'; TextList "Tool_Editor_Activated_Deactivated"; Authorization "Operate"
      ProcessValue <- "Activate_Deactivate"
      Appearance <- "Activate_Deactivate"
      on Click: InvertBit("Activate_Deactivate")
   TextField "Text field_12" at 190,593 size 335x25; Text 'Change the 100% Ration selection'
   IOField "I/O field_8" at 403,669 size 77x35; Authorization "Operate"; FormatPattern 9999.99
      ProcessValue <- "DB_MouldEditor_HMI_uData_sSelected_sPS_arFlow{1}"
      Visibility <- "DB704_MH_Value_Mixinghead{0}_AmountComponent"
      ObjectEnable <- "DB_MouldEditor_HMI_uData_sSelected_iCalculation"
      Appearance <- "DB_MouldEditor_HMI_uData_sSelected_iCalculation"
      on OnFinishInput: SetBit("DB_MouldEditor_HMI_uData_sStatusBits_xValueChanged")
   IOField "I/O field_9" at 403,703 size 77x35; Authorization "Operate"; FormatPattern 9999.99
      ProcessValue <- "DB_MouldEditor_HMI_uData_sSelected_sPS_arRatio{1}"
      Visibility <- "DB704_MH_Value_Mixinghead{0}_AmountComponent"
      Appearance <- "DB_MouldEditor_HMI_uData_sSelected_sPS_RefComponent"
      ObjectEnable <- "DB_MouldEditor_HMI_uData_sSelected_sPS_RefComponent"
      on OnFinishInput: SetBit("DB_MouldEditor_HMI_uData_sStatusBits_xValueChanged")
   IOField "I/O field_10" at 403,737 size 77x35; Authorization "Operate"; FormatPattern 9999.99
      ProcessValue <- "DB_MouldEditor_HMI_uData_sSelected_sPS_arPressure{1}"
      Visibility <- "DB704_MH_Value_Mixinghead{0}_AmountComponent"
      on OnFinishInput: SetBit("DB_MouldEditor_HMI_uData_sStatusBits_xValueChanged")
   IOField "I/O field_11" at 539,669 size 77x35; Authorization "Operate"; FormatPattern 9999.99
      ProcessValue <- "DB_MouldEditor_HMI_uData_sSelected_sPS_arFlow{2}"
      Visibility <- "DB704_MH_Value_Mixinghead{0}_AmountComponent"
      ObjectEnable <- "DB_MouldEditor_HMI_uData_sSelected_iCalculation"
      Appearance <- "DB_MouldEditor_HMI_uData_sSelected_iCalculation"
      on OnFinishInput: SetBit("DB_MouldEditor_HMI_uData_sStatusBits_xValueChanged")
   IOField "I/O field_12" at 539,703 size 77x35; Authorization "Operate"; FormatPattern 9999.99
      ProcessValue <- "DB_MouldEditor_HMI_uData_sSelected_sPS_arRatio{2}"
      Visibility <- "DB704_MH_Value_Mixinghead{0}_AmountComponent"
      Appearance <- "DB_MouldEditor_HMI_uData_sSelected_sPS_RefComponent"
      ObjectEnable <- "DB_MouldEditor_HMI_uData_sSelected_sPS_RefComponent"
      on OnFinishInput: SetBit("DB_MouldEditor_HMI_uData_sStatusBits_xValueChanged")
   IOField "I/O field_13" at 539,737 size 77x35; Authorization "Operate"; FormatPattern 9999.99
      ProcessValue <- "DB_MouldEditor_HMI_uData_sSelected_sPS_arPressure{2}"
      Visibility <- "DB704_MH_Value_Mixinghead{0}_AmountComponent"
      on OnFinishInput: SetBit("DB_MouldEditor_HMI_uData_sStatusBits_xValueChanged")
   TextField "Text field_15" at 110,669 size 236x35; Text 'Flow: [g/s]'
   TextField "Text field_16" at 110,703 size 236x35; Text 'Ratio:'
   TextField "Text field_17" at 110,737 size 236x35; Text 'Pressure:[bar]'
   Button "b_delete" at 1075,201 size 72x64; TextOff 'Delete'; PictureOff "Del"; Authorization "Operate"
      on Click: SetBit("DB_MouldEditor_HMI_uData_sStatusBits_xDeleteProgram"); "VBStore_tool_Deleted"('\Storage Card SD')
      Visibility <- "DB_MouldEditor_HMI_uData_sStatusBits_xValueChanged"
   Button "Button_3" at 326,104 size 451x32; TextOff 'Tool Editor'
   IOField "I/O field_14" at 667,143 size 185x35; Authorization "Operate"; FormatPattern ????????????????????
      ProcessValue <- "DB_MouldEditor_HMI_uData_uTools_tool_name"
      Visibility <- "DB_MouldEditor_HMI_uData_uTools_PartShot_Amount"
   Button "b_ToolAllocation" at 1075,277 size 72x64; TextOff 'Tool Alloc'; PictureOff "021-online-learning-1"
      on Click: ActivateScreen("0030_Tool Allocation", 0); SetTag("NavScreenChange", 0)
      Visibility <- "DB_MouldEditor_HMI_uData_sStatusBits_xValueChanged"
   Button "b_PartCounters" at 1075,353 size 72x64; TextOff 'Part Counter'; PictureOff "part counter"
      on Click: ActivateScreen("0887_Create Part Counter", 0); SetTag("NavScreenChange", 0)